(* Logix 5000 project; controller OWF Emulate 5570 rev 30.12; software revision 30.00; part 3 of 4 *)
(* tags used below, declared in another part *)
   OWF_Key : DINT[512,17];
(* MainProgram, continued *)

   	OWF_Key[289,15]:=338777795;
   	OWF_Key[289,16]:=945081003;
   	OWF_Key[290,13]:=1163066761;
   	OWF_Key[290,14]:=152927589;
   	OWF_Key[290,15]:=1794441803;
   	OWF_Key[290,16]:=745909431;
   	OWF_Key[291,13]:=1056792116;
   	OWF_Key[291,14]:=716761256;
   	OWF_Key[291,15]:=434777385;
   	OWF_Key[291,16]:=972035076;
   	OWF_Key[292,13]:=484357097;
   	OWF_Key[292,14]:=2101464183;
   	OWF_Key[292,15]:=1722387229;
   	OWF_Key[292,16]:=1245241283;
   	OWF_Key[293,13]:=1847549805;
   	OWF_Key[293,14]:=1256582647;
   	OWF_Key[293,15]:=854191733;
   	OWF_Key[293,16]:=1454264135;
   	OWF_Key[294,13]:=1955537619;
   	OWF_Key[294,14]:=1855656113;
   	OWF_Key[294,15]:=291670058;
   	OWF_Key[294,16]:=1334823296;
   	OWF_Key[295,13]:=429592057;
   	OWF_Key[295,14]:=2125279758;
   	OWF_Key[295,15]:=759558616;
   	OWF_Key[295,16]:=1741916674;
   	OWF_Key[296,13]:=1857086938;
   	OWF_Key[296,14]:=704728109;
   	OWF_Key[296,15]:=886421621;
   	OWF_Key[296,16]:=3201748;
   	OWF_Key[297,13]:=386252852;
   	OWF_Key[297,14]:=323092573;
   	OWF_Key[297,15]:=767083854;
   	OWF_Key[297,16]:=1353086679;
   	OWF_Key[298,13]:=1155195370;
   	OWF_Key[298,14]:=1997023534;
   	OWF_Key[298,15]:=2056641192;
   	OWF_Key[298,16]:=345689154;
   	OWF_Key[299,13]:=1620083349;
   	OWF_Key[299,14]:=211670168;
   	OWF_Key[299,15]:=811829705;
   	OWF_Key[299,16]:=277367919;
   	OWF_Key[300,13]:=1961532428;
   	OWF_Key[300,14]:=815206862;
   	OWF_Key[300,15]:=744412682;
   	OWF_Key[300,16]:=441400608;
   	OWF_Key[301,13]:=1208038755;
   	OWF_Key[301,14]:=653882227;
   	OWF_Key[301,15]:=1240796480;
   	OWF_Key[301,16]:=128162413;
   	OWF_Key[302,13]:=2049633575;
   	OWF_Key[302,14]:=1745300379;
   	OWF_Key[302,15]:=482313562;
   	OWF_Key[302,16]:=722102724;
   	OWF_Key[303,13]:=530441830;
   	OWF_Key[303,14]:=1253756416;
   	OWF_Key[303,15]:=1387935805;
   	OWF_Key[303,16]:=928482988;
   	OWF_Key[304,13]:=1989996189;
   	OWF_Key[304,14]:=86033876;
   	OWF_Key[304,15]:=488768642;
   	OWF_Key[304,16]:=1075456870;
   	OWF_Key[305,13]:=1109097795;
   	OWF_Key[305,14]:=372387132;
   	OWF_Key[305,15]:=1353015799;
   	OWF_Key[305,16]:=1061161169;
   	OWF_Key[306,13]:=783303237;
   	OWF_Key[306,14]:=1713072766;
   	OWF_Key[306,15]:=1914565908;
   	OWF_Key[306,16]:=670093717;
   	OWF_Key[307,13]:=329778336;
   	OWF_Key[307,14]:=104076356;
   	OWF_Key[307,15]:=1302500049;
   	OWF_Key[307,16]:=1142923822;
   	OWF_Key[308,13]:=1444733042;
   	OWF_Key[308,14]:=1128186410;
   	OWF_Key[308,15]:=683282754;
   	OWF_Key[308,16]:=1115169349;
   	OWF_Key[309,13]:=150257554;
   	OWF_Key[309,14]:=499012565;
   	OWF_Key[309,15]:=667227803;
   	OWF_Key[309,16]:=1601528558;
   	OWF_Key[310,13]:=580316542;
   	OWF_Key[310,14]:=276589809;
   	OWF_Key[310,15]:=319937554;
   	OWF_Key[310,16]:=1589003331;
   	OWF_Key[311,13]:=1855935330;
   	OWF_Key[311,14]:=1853361826;
   	OWF_Key[311,15]:=21601491;
   	OWF_Key[311,16]:=864859250;
   	OWF_Key[312,13]:=1594124469;
   	OWF_Key[312,14]:=432625406;
   	OWF_Key[312,15]:=295931513;
   	OWF_Key[312,16]:=1715150066;
   	OWF_Key[313,13]:=1236228216;
   	OWF_Key[313,14]:=1499623519;
   	OWF_Key[313,15]:=995144360;
   	OWF_Key[313,16]:=929655191;
   	OWF_Key[314,13]:=1016181870;
   	OWF_Key[314,14]:=1335140004;
   	OWF_Key[314,15]:=139367992;
   	OWF_Key[314,16]:=941886477;
   	OWF_Key[315,13]:=423512184;
   	OWF_Key[315,14]:=620068374;
   	OWF_Key[315,15]:=1965710084;
   	OWF_Key[315,16]:=1343328392;
   	OWF_Key[316,13]:=561716627;
   	OWF_Key[316,14]:=598814707;
   	OWF_Key[316,15]:=1265153692;
   	OWF_Key[316,16]:=316952899;
   	OWF_Key[317,13]:=112507950;
   	OWF_Key[317,14]:=319155498;
   	OWF_Key[317,15]:=961371234;
   	OWF_Key[317,16]:=593432440;
   	OWF_Key[318,13]:=1354556728;
   	OWF_Key[318,14]:=700658532;
   	OWF_Key[318,15]:=474680595;
   	OWF_Key[318,16]:=1740011842;
   	OWF_Key[319,13]:=726143028;
   	OWF_Key[319,14]:=397215194;
   	OWF_Key[319,15]:=1529304239;
   	OWF_Key[319,16]:=1797611398;
   	OWF_Key[320,13]:=800932840;
   	OWF_Key[320,14]:=197985752;
   	OWF_Key[320,15]:=1515194092;
   	OWF_Key[320,16]:=645984578;
   	OWF_Key[321,13]:=1741920313;
   	OWF_Key[321,14]:=1598171095;
   	OWF_Key[321,15]:=769783549;
   	OWF_Key[321,16]:=296019157;
   	OWF_Key[322,13]:=1307992427;
   	OWF_Key[322,14]:=648809016;
   	OWF_Key[322,15]:=2053348049;
   	OWF_Key[322,16]:=855913725;
   	OWF_Key[323,13]:=71057023;
   	OWF_Key[323,14]:=599787653;
   	OWF_Key[323,15]:=1546455656;
   	OWF_Key[323,16]:=705423056;
   	OWF_Key[324,13]:=954178807;
   	OWF_Key[324,14]:=2014078615;
   	OWF_Key[324,15]:=1878645210;
   	OWF_Key[324,16]:=856338194;
   	OWF_Key[325,13]:=1706921177;
   	OWF_Key[325,14]:=483825803;
   	OWF_Key[325,15]:=983348168;
   	OWF_Key[325,16]:=1208835096;
   	OWF_Key[326,13]:=1598778839;
   	OWF_Key[326,14]:=1893467300;
   	OWF_Key[326,15]:=580814559;
   	OWF_Key[326,16]:=2131522844;
   	OWF_Key[327,13]:=244599566;
   	OWF_Key[327,14]:=555308622;
   	OWF_Key[327,15]:=1516006940;
   	OWF_Key[327,16]:=1173694990;
   	OWF_Key[328,13]:=941443323;
   	OWF_Key[328,14]:=843686349;
   	OWF_Key[328,15]:=1922095669;
   	OWF_Key[328,16]:=1779289712;
   	OWF_Key[329,13]:=1304931617;
   	OWF_Key[329,14]:=1151000137;
   	OWF_Key[329,15]:=124471029;
   	OWF_Key[329,16]:=1971689967;
   	OWF_Key[330,13]:=1453682887;
   	OWF_Key[330,14]:=805069671;
   	OWF_Key[330,15]:=1650012438;
   	OWF_Key[330,16]:=1453746600;
   	OWF_Key[331,13]:=590923085;
   	OWF_Key[331,14]:=1002744768;
   	OWF_Key[331,15]:=1426998178;
   	OWF_Key[331,16]:=821237014;
   	OWF_Key[332,13]:=1614486384;
   	OWF_Key[332,14]:=2104870625;
   	OWF_Key[332,15]:=315969258;
   	OWF_Key[332,16]:=1578924085;
   	OWF_Key[333,13]:=2041706571;
   	OWF_Key[333,14]:=16774744;
   	OWF_Key[333,15]:=915382048;
   	OWF_Key[333,16]:=648804525;
   	OWF_Key[334,13]:=316000875;
   	OWF_Key[334,14]:=1862306372;
   	OWF_Key[334,15]:=1355759476;
   	OWF_Key[334,16]:=1859145934;
   	OWF_Key[335,13]:=1975045396;
   	OWF_Key[335,14]:=327165606;
   	OWF_Key[335,15]:=834469435;
   	OWF_Key[335,16]:=1485936747;
   	OWF_Key[336,13]:=1461136409;
   	OWF_Key[336,14]:=278026422;
   	OWF_Key[336,15]:=1210238525;
   	OWF_Key[336,16]:=405251428;
   	OWF_Key[337,13]:=1643706608;
   	OWF_Key[337,14]:=1161448288;
   	OWF_Key[337,15]:=51875454;
   	OWF_Key[337,16]:=1551504033;
   	OWF_Key[338,13]:=1459047679;
   	OWF_Key[338,14]:=1308895253;
   	OWF_Key[338,15]:=1148280820;
   	OWF_Key[338,16]:=1216977140;
   	OWF_Key[339,13]:=829366181;
   	OWF_Key[339,14]:=840670868;
   	OWF_Key[339,15]:=2100768505;
   	OWF_Key[339,16]:=509465283;
   	OWF_Key[340,13]:=10547943;
   	OWF_Key[340,14]:=649144044;
   	OWF_Key[340,15]:=919338342;
   	OWF_Key[340,16]:=1030770615;
   	OWF_Key[341,13]:=1793689517;
   	OWF_Key[341,14]:=161281212;
   	OWF_Key[341,15]:=535831803;
   	OWF_Key[341,16]:=208840162;
   	OWF_Key[342,13]:=199305394;
   	OWF_Key[342,14]:=792165041;
   	OWF_Key[342,15]:=1982050062;
   	OWF_Key[342,16]:=590342057;
   	OWF_Key[343,13]:=2112922264;
   	OWF_Key[343,14]:=1923655750;
   	OWF_Key[343,15]:=988358550;
   	OWF_Key[343,16]:=257463890;
   	OWF_Key[344,13]:=1265962317;
   	OWF_Key[344,14]:=705872158;
   	OWF_Key[344,15]:=1873115819;
   	OWF_Key[344,16]:=1158681719;
   	OWF_Key[345,13]:=365212730;
   	OWF_Key[345,14]:=1387331228;
   	OWF_Key[345,15]:=1953063521;
   	OWF_Key[345,16]:=190819161;
   	OWF_Key[346,13]:=1487999543;
   	OWF_Key[346,14]:=213890483;
   	OWF_Key[346,15]:=2033855619;
   	OWF_Key[346,16]:=1750025558;
   	OWF_Key[347,13]:=1214378656;
   	OWF_Key[347,14]:=1204880672;
   	OWF_Key[347,15]:=1632730149;
   	OWF_Key[347,16]:=1524207983;
   	OWF_Key[348,13]:=505673370;
   	OWF_Key[348,14]:=584281114;
   	OWF_Key[348,15]:=1062156090;
   	OWF_Key[348,16]:=1569692077;
   	OWF_Key[349,13]:=575514820;
   	OWF_Key[349,14]:=286269877;
   	OWF_Key[349,15]:=1401152444;
   	OWF_Key[349,16]:=392054891;
   	OWF_Key[350,13]:=1748777147;
   	OWF_Key[350,14]:=2083193089;
   	OWF_Key[350,15]:=1572988760;
   	OWF_Key[350,16]:=2138728050;
   	OWF_Key[351,13]:=1202747954;
   	OWF_Key[351,14]:=820441372;
   	OWF_Key[351,15]:=1077683802;
   	OWF_Key[351,16]:=1924437405;
   	OWF_Key[352,13]:=2014139620;
   	OWF_Key[352,14]:=1335552778;
   	OWF_Key[352,15]:=775142346;
   	OWF_Key[352,16]:=1227681831;
   	OWF_Key[353,13]:=48430552;
   	OWF_Key[353,14]:=1049121167;
   	OWF_Key[353,15]:=287349008;
   	OWF_Key[353,16]:=684937982;
   	OWF_Key[354,13]:=214282945;
   	OWF_Key[354,14]:=1789370232;
   	OWF_Key[354,15]:=1634651577;
   	OWF_Key[354,16]:=1956112331;
   	OWF_Key[355,13]:=672289927;
   	OWF_Key[355,14]:=1636493386;
   	OWF_Key[355,15]:=335595154;
   	OWF_Key[355,16]:=1103131647;
   	OWF_Key[356,13]:=1665909380;
   	OWF_Key[356,14]:=940971670;
   	OWF_Key[356,15]:=1085160366;
   	OWF_Key[356,16]:=793143189;
   	OWF_Key[357,13]:=2119272361;
   	OWF_Key[357,14]:=887959070;
   	OWF_Key[357,15]:=1660665421;
   	OWF_Key[357,16]:=11136188;
   	OWF_Key[358,13]:=104486906;
   	OWF_Key[358,14]:=2089719193;
   	OWF_Key[358,15]:=694497781;
   	OWF_Key[358,16]:=1060026839;
   	OWF_Key[359,13]:=1242387453;
   	OWF_Key[359,14]:=265858260;
   	OWF_Key[359,15]:=2122202457;
   	OWF_Key[359,16]:=1166357817;
   	OWF_Key[360,13]:=1891573758;
   	OWF_Key[360,14]:=260897043;
   	OWF_Key[360,15]:=802879836;
   	OWF_Key[360,16]:=1234754780;
   	OWF_Key[361,13]:=1348865357;
   	OWF_Key[361,14]:=832359419;
   	OWF_Key[361,15]:=845448176;
   	OWF_Key[361,16]:=1220047530;
   	OWF_Key[362,13]:=1270006551;
   	OWF_Key[362,14]:=1384711650;
   	OWF_Key[362,15]:=1730649878;
   	OWF_Key[362,16]:=1662691495;
   	OWF_Key[363,13]:=1752061486;
   	OWF_Key[363,14]:=1230806191;
   	OWF_Key[363,15]:=1489100239;
   	OWF_Key[363,16]:=1531443934;
   	OWF_Key[364,13]:=2101981980;
   	OWF_Key[364,14]:=1458680843;
   	OWF_Key[364,15]:=1859987205;
   	OWF_Key[364,16]:=1123074689;
   	OWF_Key[365,13]:=1302345128;
   	OWF_Key[365,14]:=1781711563;
   	OWF_Key[365,15]:=782583437;
   	OWF_Key[365,16]:=1751869154;
   	OWF_Key[366,13]:=1269026032;
   	OWF_Key[366,14]:=1565939600;
   	OWF_Key[366,15]:=796422412;
   	OWF_Key[366,16]:=1413232287;
   	OWF_Key[367,13]:=994794909;
   	OWF_Key[367,14]:=940478114;
   	OWF_Key[367,15]:=1927914407;
   	OWF_Key[367,16]:=516452424;
   	OWF_Key[368,13]:=353288391;
   	OWF_Key[368,14]:=1006705053;
   	OWF_Key[368,15]:=833926143;
   	OWF_Key[368,16]:=1833767657;
   	OWF_Key[369,13]:=830407689;
   	OWF_Key[369,14]:=1883974526;
   	OWF_Key[369,15]:=32397573;
   	OWF_Key[369,16]:=1610932340;
   	OWF_Key[370,13]:=1570129652;
   	OWF_Key[370,14]:=2060232729;
   	OWF_Key[370,15]:=1139326171;
   	OWF_Key[370,16]:=1746459602;
   	OWF_Key[371,13]:=1872850139;
   	OWF_Key[371,14]:=1311501626;
   	OWF_Key[371,15]:=1382272678;
   	OWF_Key[371,16]:=2011320514;
   	OWF_Key[372,13]:=1045068510;
   	OWF_Key[372,14]:=393024892;
   	OWF_Key[372,15]:=634135353;
   	OWF_Key[372,16]:=1470069055;
   	OWF_Key[373,13]:=328609956;
   	OWF_Key[373,14]:=1383192207;
   	OWF_Key[373,15]:=1535515614;
   	OWF_Key[373,16]:=715297357;
   	OWF_Key[374,13]:=620723337;
   	OWF_Key[374,14]:=454533633;
   	OWF_Key[374,15]:=658920899;
   	OWF_Key[374,16]:=1672648486;
   	OWF_Key[375,13]:=229075100;
   	OWF_Key[375,14]:=599980880;
   	OWF_Key[375,15]:=2120266548;
   	OWF_Key[375,16]:=1605768993;
   	OWF_Key[376,13]:=434021335;
   	OWF_Key[376,14]:=785720651;
   	OWF_Key[376,15]:=2060675124;
   	OWF_Key[376,16]:=1067843577;
   	OWF_Key[377,13]:=1864505716;
   	OWF_Key[377,14]:=434694751;
   	OWF_Key[377,15]:=2090811;
   	OWF_Key[377,16]:=2088506733;
   	OWF_Key[378,13]:=709750540;
   	OWF_Key[378,14]:=1972107009;
   	OWF_Key[378,15]:=241297992;
   	OWF_Key[378,16]:=1837533029;
   	OWF_Key[379,13]:=522199474;
   	OWF_Key[379,14]:=1365297600;
   	OWF_Key[379,15]:=315087364;
   	OWF_Key[379,16]:=1676043165;
   	OWF_Key[380,13]:=1339113249;
   	OWF_Key[380,14]:=1694379432;
   	OWF_Key[380,15]:=291694756;
   	OWF_Key[380,16]:=265747760;
   	OWF_Key[381,13]:=552624291;
   	OWF_Key[381,14]:=1165273822;
   	OWF_Key[381,15]:=1794394231;
   	OWF_Key[381,16]:=736035571;
   	OWF_Key[382,13]:=715064081;
   	OWF_Key[382,14]:=1125061568;
   	OWF_Key[382,15]:=77469684;
   	OWF_Key[382,16]:=2053028533;
   	OWF_Key[383,13]:=1153340465;
   	OWF_Key[383,14]:=408686771;
   	OWF_Key[383,15]:=1420990686;
   	OWF_Key[383,16]:=1762240643;
   	OWF_Key[384,0]:=1123644528;
   	OWF_Key[384,1]:=327294325;
   	OWF_Key[384,2]:=89446114;
   	OWF_Key[384,3]:=400023116;
   	OWF_Key[384,4]:=2133600475;
   	OWF_Key[384,5]:=1972870607;
   	OWF_Key[384,6]:=1960923513;
   	OWF_Key[384,7]:=1610917558;
   	OWF_Key[384,8]:=1384593970;
   	OWF_Key[384,9]:=478162938;
   	OWF_Key[384,10]:=482847716;
   	OWF_Key[384,11]:=105738552;
   	OWF_Key[384,12]:=1816536681;
   	OWF_Key[384,13]:=1691613707;
   	OWF_Key[384,14]:=402827396;
   	OWF_Key[384,15]:=933136802;
   	OWF_Key[384,16]:=200058548;
   	OWF_Key[385,0]:=1190356074;
   	OWF_Key[385,1]:=1735118759;
   	OWF_Key[385,2]:=534327591;
   	OWF_Key[385,3]:=1988815940;
   	OWF_Key[385,4]:=2109121553;
   	OWF_Key[385,5]:=1649017839;
   	OWF_Key[385,6]:=1489916775;
   	OWF_Key[385,7]:=1296815713;
   	OWF_Key[385,8]:=64645432;
   	OWF_Key[385,9]:=1103622136;
   	OWF_Key[385,10]:=673381504;
   	OWF_Key[385,11]:=453919901;
   	OWF_Key[385,12]:=240114348;
   	OWF_Key[385,13]:=1623339818;
   	OWF_Key[385,14]:=634006860;
   	OWF_Key[385,15]:=427414237;
   	OWF_Key[385,16]:=118494102;
   	OWF_Key[386,0]:=15965030;
   	OWF_Key[386,1]:=1184331497;
   	OWF_Key[386,2]:=176506727;
   	OWF_Key[386,3]:=600317579;
   	OWF_Key[386,4]:=760943662;
   	OWF_Key[386,5]:=1416388614;
   	OWF_Key[386,6]:=579063372;
   	OWF_Key[386,7]:=193484260;
   	OWF_Key[386,8]:=886558396;
   	OWF_Key[386,9]:=1929832978;
   	OWF_Key[386,10]:=1586193234;
   	OWF_Key[386,11]:=1446931923;
   	OWF_Key[386,12]:=443040518;
   	OWF_Key[386,13]:=1789561753;
   	OWF_Key[386,14]:=812617742;
   	OWF_Key[386,15]:=1005140005;
   	OWF_Key[386,16]:=1763651041;
   	OWF_Key[387,0]:=473065605;
   	OWF_Key[387,1]:=1971577610;
   	OWF_Key[387,2]:=1382360800;
   	OWF_Key[387,3]:=668173573;
   	OWF_Key[387,4]:=1949911116;
   	OWF_Key[387,5]:=699197275;
   	OWF_Key[387,6]:=1386638121;
   	OWF_Key[387,7]:=1668072067;
   	OWF_Key[387,8]:=1597740321;
   	OWF_Key[387,9]:=588219297;
   	OWF_Key[387,10]:=107304456;
   	OWF_Key[387,11]:=1679213174;
   	OWF_Key[387,12]:=1164872061;
   	OWF_Key[387,13]:=2134830521;
   	OWF_Key[387,14]:=938176584;
   	OWF_Key[387,15]:=350011980;
   	OWF_Key[387,16]:=1306194849;
   	OWF_Key[388,0]:=1219015982;
   	OWF_Key[388,1]:=1110225865;
   	OWF_Key[388,2]:=525391525;
   	OWF_Key[388,3]:=1016867921;
   	OWF_Key[388,4]:=388802829;
   	OWF_Key[388,5]:=809856191;
   	OWF_Key[388,6]:=1220410729;
   	OWF_Key[388,7]:=566369721;
   	OWF_Key[388,8]:=971805674;
   	OWF_Key[388,9]:=1369966763;
   	OWF_Key[388,10]:=897986535;
   	OWF_Key[388,11]:=683802913;
   	OWF_Key[388,12]:=454325621;
   	OWF_Key[388,13]:=1811777432;
   	OWF_Key[388,14]:=1096785551;
   	OWF_Key[388,15]:=1387324969;
   	OWF_Key[388,16]:=2144832821;
   	OWF_Key[389,0]:=1732712476;
   	OWF_Key[389,1]:=2117139316;
   	OWF_Key[389,2]:=1006496162;
   	OWF_Key[389,3]:=1856826815;
   	OWF_Key[389,4]:=314563872;
   	OWF_Key[389,5]:=1436637226;
   	OWF_Key[389,6]:=829596455;
   	OWF_Key[389,7]:=1658267507;
   	OWF_Key[389,8]:=1423018056;
   	OWF_Key[389,9]:=403040411;
   	OWF_Key[389,10]:=1702067466;
   	OWF_Key[389,11]:=424286356;
   	OWF_Key[389,12]:=1660115278;
   	OWF_Key[389,13]:=665344609;
   	OWF_Key[389,14]:=780639910;
   	OWF_Key[389,15]:=501642388;
   	OWF_Key[389,16]:=959856039;
   	OWF_Key[390,0]:=629397116;
   	OWF_Key[390,1]:=2100981858;
   	OWF_Key[390,2]:=959457952;
   	OWF_Key[390,3]:=344681006;
   	OWF_Key[390,4]:=2055412444;
   	OWF_Key[390,5]:=890642893;
   	OWF_Key[390,6]:=920375373;
   	OWF_Key[390,7]:=1537083478;
   	OWF_Key[390,8]:=553468104;
   	OWF_Key[390,9]:=344155898;
   	OWF_Key[390,10]:=117485162;
   	OWF_Key[390,11]:=1653582078;
   	OWF_Key[390,12]:=1911913238;
   	OWF_Key[390,13]:=1399825354;
   	OWF_Key[390,14]:=1201110775;
   	OWF_Key[390,15]:=1363257890;
   	OWF_Key[390,16]:=299268868;
   	OWF_Key[391,0]:=704460495;
   	OWF_Key[391,1]:=2095392130;
   	OWF_Key[391,2]:=1380916171;
   	OWF_Key[391,3]:=1505402993;
   	OWF_Key[391,4]:=1762832652;
   	OWF_Key[391,5]:=1819207163;
   	OWF_Key[391,6]:=1230495993;
   	OWF_Key[391,7]:=175012694;
   	OWF_Key[391,8]:=497472778;
   	OWF_Key[391,9]:=1117394135;
   	OWF_Key[391,10]:=1939865321;
   	OWF_Key[391,11]:=1263415657;
   	OWF_Key[391,12]:=1025065602;
   	OWF_Key[391,13]:=1967755854;
   	OWF_Key[391,14]:=332938538;
   	OWF_Key[391,15]:=198300463;
   	OWF_Key[391,16]:=654647784;
   	OWF_Key[392,0]:=1877447257;
   	OWF_Key[392,1]:=1406678132;
   	OWF_Key[392,2]:=2092744173;
   	OWF_Key[392,3]:=769562260;
   	OWF_Key[392,4]:=332946273;
   	OWF_Key[392,5]:=1266561390;
   	OWF_Key[392,6]:=2067638902;
   	OWF_Key[392,7]:=931566009;
   	OWF_Key[392,8]:=769768789;
   	OWF_Key[392,9]:=409067196;
   	OWF_Key[392,10]:=50536829;
   	OWF_Key[392,11]:=1292364619;
   	OWF_Key[392,12]:=670226040;
   	OWF_Key[392,13]:=1703281565;
   	OWF_Key[392,14]:=1817010827;
   	OWF_Key[392,15]:=471741373;
   	OWF_Key[392,16]:=2110439650;
   	OWF_Key[393,0]:=558191637;
   	OWF_Key[393,1]:=189579802;
   	OWF_Key[393,2]:=70773707;
   	OWF_Key[393,3]:=1198325196;
   	OWF_Key[393,4]:=896109359;
   	OWF_Key[393,5]:=844755332;
   	OWF_Key[393,6]:=1694894433;
   	OWF_Key[393,7]:=1727275555;
   	OWF_Key[393,8]:=1153084870;
   	OWF_Key[393,9]:=1296582337;
   	OWF_Key[393,10]:=395365370;
   	OWF_Key[393,11]:=2067650742;
   	OWF_Key[393,12]:=537962770;
   	OWF_Key[393,13]:=875213948;
   	OWF_Key[393,14]:=1879930164;
   	OWF_Key[393,15]:=215274890;
   	OWF_Key[393,16]:=765449581;
   	OWF_Key[394,0]:=1209351764;
   	OWF_Key[394,1]:=1929455118;
   	OWF_Key[394,2]:=1364106375;
   	OWF_Key[394,3]:=1935297266;
   	OWF_Key[394,4]:=735170043;
   	OWF_Key[394,5]:=651296485;
   	OWF_Key[394,6]:=617760457;
   	OWF_Key[394,7]:=781979719;
   	OWF_Key[394,8]:=646465543;
   	OWF_Key[394,9]:=1306700206;
   	OWF_Key[394,10]:=293993545;
   	OWF_Key[394,11]:=1718622122;
   	OWF_Key[394,12]:=1921118428;
   	OWF_Key[394,13]:=1626271946;
   	OWF_Key[394,14]:=755823439;
   	OWF_Key[394,15]:=1641210106;
   	OWF_Key[394,16]:=1161503765;
   	OWF_Key[395,0]:=1612949080;
   	OWF_Key[395,1]:=37057564;
   	OWF_Key[395,2]:=969908110;
   	OWF_Key[395,3]:=325860815;
   	OWF_Key[395,4]:=1977473562;
   	OWF_Key[395,5]:=1574820053;
   	OWF_Key[395,6]:=1865550696;
   	OWF_Key[395,7]:=57204164;
   	OWF_Key[395,8]:=1719255575;
   	OWF_Key[395,9]:=987103474;
   	OWF_Key[395,10]:=1664178903;
   	OWF_Key[395,11]:=1419145457;
   	OWF_Key[395,12]:=823480756;
   	OWF_Key[395,13]:=572322380;
   	OWF_Key[395,14]:=1278186542;
   	OWF_Key[395,15]:=1398628562;
   	OWF_Key[395,16]:=960886128;
   	OWF_Key[396,0]:=880749436;
   	OWF_Key[396,1]:=605599712;
   	OWF_Key[396,2]:=222767252;
   	OWF_Key[396,3]:=1351229525;
   	OWF_Key[396,4]:=965055471;
   	OWF_Key[396,5]:=2131021532;
   	OWF_Key[396,6]:=1801157192;
   	OWF_Key[396,7]:=1328575616;
   	OWF_Key[396,8]:=1729664556;
   	OWF_Key[396,9]:=1541266684;
   	OWF_Key[396,10]:=1930731347;
   	OWF_Key[396,11]:=636772215;
   	OWF_Key[396,12]:=579829843;
   	OWF_Key[396,13]:=1501270875;
   	OWF_Key[396,14]:=1149353205;
   	OWF_Key[396,15]:=808254363;
   	OWF_Key[396,16]:=988338201;
   	OWF_Key[397,0]:=624471172;
   	OWF_Key[397,1]:=1693671742;
   	OWF_Key[397,2]:=489913198;
   	OWF_Key[397,3]:=1222896940;
   	OWF_Key[397,4]:=839749689;
   	OWF_Key[397,5]:=1565229034;
   	OWF_Key[397,6]:=1344903047;
   	OWF_Key[397,7]:=1571644055;
   	OWF_Key[397,8]:=781586711;
   	OWF_Key[397,9]:=13493181;
   	OWF_Key[397,10]:=1927637652;
   	OWF_Key[397,11]:=1995483867;
   	OWF_Key[397,12]:=1669800219;
   	OWF_Key[397,13]:=176222652;
   	OWF_Key[397,14]:=1637048009;
   	OWF_Key[397,15]:=2111318472;
   	OWF_Key[397,16]:=1461920624;
   	OWF_Key[398,0]:=1783356394;
   	OWF_Key[398,1]:=467500457;
   	OWF_Key[398,2]:=1812456881;
   	OWF_Key[398,3]:=474627191;
   	OWF_Key[398,4]:=1591060643;
   	OWF_Key[398,5]:=1161312513;
   	OWF_Key[398,6]:=1197289822;
   	OWF_Key[398,7]:=1616351944;
   	OWF_Key[398,8]:=242758526;
   	OWF_Key[398,9]:=1905091041;
   	OWF_Key[398,10]:=1660565429;
   	OWF_Key[398,11]:=1870317022;
   	OWF_Key[398,12]:=431717124;
   	OWF_Key[398,13]:=1882304375;
   	OWF_Key[398,14]:=145069520;
   	OWF_Key[398,15]:=364490524;
   	OWF_Key[398,16]:=1557624578;
   	OWF_Key[399,0]:=1469797541;
   	OWF_Key[399,1]:=1311253024;
   	OWF_Key[399,2]:=1349819562;
   	OWF_Key[399,3]:=1218316421;
   	OWF_Key[399,4]:=595675644;
   	OWF_Key[399,5]:=503087038;
   	OWF_Key[399,6]:=884474462;
   	OWF_Key[399,7]:=1474946218;
   	OWF_Key[399,8]:=267390419;
   	OWF_Key[399,9]:=243266912;
   	OWF_Key[399,10]:=379115072;
   	OWF_Key[399,11]:=1550234120;
   	OWF_Key[399,12]:=1290918739;
   	OWF_Key[399,13]:=660998652;
   	OWF_Key[399,14]:=1858734974;
   	OWF_Key[399,15]:=1056569339;
   	OWF_Key[399,16]:=1220610346;
   	OWF_Key[400,0]:=426350853;
   	OWF_Key[400,1]:=1457837182;
   	OWF_Key[400,2]:=1472791955;
   	OWF_Key[400,3]:=594242150;
   	OWF_Key[400,4]:=986024935;
   	OWF_Key[400,5]:=2045216485;
   	OWF_Key[400,6]:=547495341;
   	OWF_Key[400,7]:=1307195620;
   	OWF_Key[400,8]:=1910496756;
   	OWF_Key[400,9]:=1998696686;
   	OWF_Key[400,10]:=2136331173;
   	OWF_Key[400,11]:=107427988;
   	OWF_Key[400,12]:=816643110;
   	OWF_Key[400,13]:=1027059949;
   	OWF_Key[400,14]:=1065404919;
   	OWF_Key[400,15]:=137059426;
   	OWF_Key[400,16]:=2016380687;
   	OWF_Key[401,0]:=1275943308;
   	OWF_Key[401,1]:=1051704736;
   	OWF_Key[401,2]:=178716534;
   	OWF_Key[401,3]:=240880497;
   	OWF_Key[401,4]:=858624779;
   	OWF_Key[401,5]:=200115622;
   	OWF_Key[401,6]:=1420797872;
   	OWF_Key[401,7]:=1915747964;
   	OWF_Key[401,8]:=773670025;
   	OWF_Key[401,9]:=62218432;
   	OWF_Key[401,10]:=2062058736;
   	OWF_Key[401,11]:=464986808;
   	OWF_Key[401,12]:=1797617676;
   	OWF_Key[401,13]:=27012266;
   	OWF_Key[401,14]:=1795140434;
   	OWF_Key[401,15]:=1870046730;
   	OWF_Key[401,16]:=1213756716;
   	OWF_Key[402,0]:=635400718;
   	OWF_Key[402,1]:=602499652;
   	OWF_Key[402,2]:=547615363;
   	OWF_Key[402,3]:=433431976;
   	OWF_Key[402,4]:=212181673;
   	OWF_Key[402,5]:=436292151;
   	OWF_Key[402,6]:=713149480;
   	OWF_Key[402,7]:=791790870;
   	OWF_Key[402,8]:=930542692;
   	OWF_Key[402,9]:=347398757;
   	OWF_Key[402,10]:=1486676141;
   	OWF_Key[402,11]:=1295870258;
   	OWF_Key[402,12]:=1800259834;
   	OWF_Key[402,13]:=414928284;
   	OWF_Key[402,14]:=1194374331;
   	OWF_Key[402,15]:=1088052810;
   	OWF_Key[402,16]:=1505009395;
   	OWF_Key[403,0]:=985408697;
   	OWF_Key[403,1]:=58290271;
   	OWF_Key[403,2]:=649996824;
   	OWF_Key[403,3]:=87207318;
   	OWF_Key[403,4]:=1732847835;
   	OWF_Key[403,5]:=1381921644;
   	OWF_Key[403,6]:=1946940514;
   	OWF_Key[403,7]:=2069056016;
   	OWF_Key[403,8]:=65792540;
   	OWF_Key[403,9]:=1178411609;
   	OWF_Key[403,10]:=1663226500;
   	OWF_Key[403,11]:=453326667;
   	OWF_Key[403,12]:=220588916;
   	OWF_Key[403,13]:=1526064465;
   	OWF_Key[403,14]:=455636350;
   	OWF_Key[403,15]:=1683363899;
   	OWF_Key[403,16]:=2046796746;
   	OWF_Key[404,0]:=737681872;
   	OWF_Key[404,1]:=1866742463;
   	OWF_Key[404,2]:=434437596;
   	OWF_Key[404,3]:=1666265441;
   	OWF_Key[404,4]:=837265743;
   	OWF_Key[404,5]:=1571357242;
   	OWF_Key[404,6]:=1309709069;
   	OWF_Key[404,7]:=1932232725;
   	OWF_Key[404,8]:=863118724;
   	OWF_Key[404,9]:=667703742;
   	OWF_Key[404,10]:=1352555970;
   	OWF_Key[404,11]:=1506316314;
   	OWF_Key[404,12]:=264070247;
   	OWF_Key[404,13]:=1445468590;
   	OWF_Key[404,14]:=1972588571;
   	OWF_Key[404,15]:=155474394;
   	OWF_Key[404,16]:=1723592618;
   	OWF_Key[405,0]:=535700331;
   	OWF_Key[405,1]:=1966380749;
   	OWF_Key[405,2]:=684673087;
   	OWF_Key[405,3]:=45426188;
   	OWF_Key[405,4]:=1145115607;
   	OWF_Key[405,5]:=1242157266;
   	OWF_Key[405,6]:=934650184;
   	OWF_Key[405,7]:=426034024;
   	OWF_Key[405,8]:=819715969;
   	OWF_Key[405,9]:=1147277411;
   	OWF_Key[405,10]:=1076796787;
   	OWF_Key[405,11]:=1088154061;
   	OWF_Key[405,12]:=1076643300;
   	OWF_Key[405,13]:=901250297;
   	OWF_Key[405,14]:=1832803426;
   	OWF_Key[405,15]:=1119995119;
   	OWF_Key[405,16]:=678607113;
   	OWF_Key[406,0]:=1617337029;
   	OWF_Key[406,1]:=159618416;
   	OWF_Key[406,2]:=1508617393;
   	OWF_Key[406,3]:=1335810724;
   	OWF_Key[406,4]:=1187713919;
   	OWF_Key[406,5]:=1229364024;
   	OWF_Key[406,6]:=1698030676;
   	OWF_Key[406,7]:=513154543;
   	OWF_Key[406,8]:=367641541;
   	OWF_Key[406,9]:=840136748;
   	OWF_Key[406,10]:=260274723;
   	OWF_Key[406,11]:=1687968394;
   	OWF_Key[406,12]:=1955395556;
   	OWF_Key[406,13]:=1564767792;
   	OWF_Key[406,14]:=113027328;
   	OWF_Key[406,15]:=697237787;
   	OWF_Key[406,16]:=1612309181;
   	OWF_Key[407,0]:=1876867906;
   	OWF_Key[407,1]:=1611698278;
   	OWF_Key[407,2]:=776016439;
   	OWF_Key[407,3]:=509525515;
   	OWF_Key[407,4]:=1519736046;
   	OWF_Key[407,5]:=728378544;
   	OWF_Key[407,6]:=1416880690;
   	OWF_Key[407,7]:=666194178;
   	OWF_Key[407,8]:=751167067;
   	OWF_Key[407,9]:=1601561182;
   	OWF_Key[407,10]:=917046526;
   	OWF_Key[407,11]:=760269565;
   	OWF_Key[407,12]:=1644678903;
   	OWF_Key[407,13]:=2108054212;
   	OWF_Key[407,14]:=2076036808;
   	OWF_Key[407,15]:=1696466385;
   	OWF_Key[407,16]:=436140396;
   	OWF_Key[408,0]:=1035116191;
   	OWF_Key[408,1]:=1894535674;
   	OWF_Key[408,2]:=97626570;
   	OWF_Key[408,3]:=552482263;
   	OWF_Key[408,4]:=2020766682;
   	OWF_Key[408,5]:=1294987990;
   	OWF_Key[408,6]:=1547272803;
   	OWF_Key[408,7]:=335685718;
   	OWF_Key[408,8]:=1767084616;
   	OWF_Key[408,9]:=51037054;
   	OWF_Key[408,10]:=134869686;
   	OWF_Key[408,11]:=436500898;
   	OWF_Key[408,12]:=1555893409;
   	OWF_Key[408,13]:=1652214910;
   	OWF_Key[408,14]:=1803890040;
   	OWF_Key[408,15]:=350021584;
   	OWF_Key[408,16]:=918818858;
   	OWF_Key[409,0]:=2084739708;
   	OWF_Key[409,1]:=921373142;
   	OWF_Key[409,2]:=164942549;
   	OWF_Key[409,3]:=1720778444;
   	OWF_Key[409,4]:=960484409;
   	OWF_Key[409,5]:=1618501736;
   	OWF_Key[409,6]:=530958119;
   	OWF_Key[409,7]:=848389038;
   	OWF_Key[409,8]:=391885234;
   	OWF_Key[409,9]:=71564478;
   	OWF_Key[409,10]:=1531808560;
   	OWF_Key[409,11]:=2034827564;
   	OWF_Key[409,12]:=841819950;
   	OWF_Key[409,13]:=1684975312;
   	OWF_Key[409,14]:=2127333534;
   	OWF_Key[409,15]:=1974249562;
   	OWF_Key[409,16]:=1136773476;
   	OWF_Key[410,0]:=1340202885;
   	OWF_Key[410,1]:=2146847724;
   	OWF_Key[410,2]:=1265909703;
   	OWF_Key[410,3]:=835259095;
   	OWF_Key[410,4]:=996599140;
   	OWF_Key[410,5]:=1402108171;
   	OWF_Key[410,6]:=296651482;
   	OWF_Key[410,7]:=1424983826;
   	OWF_Key[410,8]:=419634320;
   	OWF_Key[410,9]:=877068425;
   	OWF_Key[410,10]:=1381222120;
   	OWF_Key[410,11]:=1915385144;
   	OWF_Key[410,12]:=1650543850;
   	OWF_Key[410,13]:=1745372635;
   	OWF_Key[410,14]:=2079645439;
   	OWF_Key[410,15]:=1804225655;
   	OWF_Key[410,16]:=1540427086;
   	OWF_Key[411,0]:=1018418210;
   	OWF_Key[411,1]:=6832204;
   	OWF_Key[411,2]:=140201042;
   	OWF_Key[411,3]:=833534206;
   	OWF_Key[411,4]:=1656655246;
   	OWF_Key[411,5]:=2040220336;
   	OWF_Key[411,6]:=2065264367;
   	OWF_Key[411,7]:=2395885;
   	OWF_Key[411,8]:=2081052196;
   	OWF_Key[411,9]:=685196918;
   	OWF_Key[411,10]:=211981018;
   	OWF_Key[411,11]:=1920575130;
   	OWF_Key[411,12]:=525356832;
   	OWF_Key[411,13]:=1161758941;
   	OWF_Key[411,14]:=166651162;
   	OWF_Key[411,15]:=334734559;
   	OWF_Key[411,16]:=12647565;
   	OWF_Key[412,0]:=1473284706;
   	OWF_Key[412,1]:=1689237493;
   	OWF_Key[412,2]:=227217910;
   	OWF_Key[412,3]:=125487887;
   	OWF_Key[412,4]:=963863316;
   	OWF_Key[412,5]:=1586790226;
   	OWF_Key[412,6]:=1690936455;
   	OWF_Key[412,7]:=1248985432;
   	OWF_Key[412,8]:=857799518;
   	OWF_Key[412,9]:=1801132884;
   	OWF_Key[412,10]:=1364107014;
   	OWF_Key[412,11]:=1356990110;
   	OWF_Key[412,12]:=49851296;
   	OWF_Key[412,13]:=1896029743;
   	OWF_Key[412,14]:=168052664;
   	OWF_Key[412,15]:=1559863538;
   	OWF_Key[412,16]:=868031175;
   	OWF_Key[413,0]:=973211649;
   	OWF_Key[413,1]:=1156672633;
   	OWF_Key[413,2]:=666204571;
   	OWF_Key[413,3]:=1164315747;
   	OWF_Key[413,4]:=909812080;
   	OWF_Key[413,5]:=665362095;
   	OWF_Key[413,6]:=1859789997;
   	OWF_Key[413,7]:=57252400;
   	OWF_Key[413,8]:=450810821;
   	OWF_Key[413,9]:=745456181;
   	OWF_Key[413,10]:=1817188413;
   	OWF_Key[413,11]:=2016658328;
   	OWF_Key[413,12]:=1512212636;
   	OWF_Key[413,13]:=129954824;
   	OWF_Key[413,14]:=2044212889;
   	OWF_Key[413,15]:=834946124;
   	OWF_Key[413,16]:=602936897;
   	OWF_Key[414,0]:=113894710;
   	OWF_Key[414,1]:=242368547;
   	OWF_Key[414,2]:=651374774;
   	OWF_Key[414,3]:=27204543;
   	OWF_Key[414,4]:=318834520;
   	OWF_Key[414,5]:=1846049833;
   	OWF_Key[414,6]:=1549322185;
   	OWF_Key[414,7]:=1586245847;
   	OWF_Key[414,8]:=1660644610;
   	OWF_Key[414,9]:=671591771;
   	OWF_Key[414,10]:=463573;
   	OWF_Key[414,11]:=699541753;
   	OWF_Key[414,12]:=243773552;
   	OWF_Key[414,13]:=273956214;
   	OWF_Key[414,14]:=1999906248;
   	OWF_Key[414,15]:=1432020015;
   	OWF_Key[414,16]:=1459843515;
   	OWF_Key[415,0]:=1764109547;
   	OWF_Key[415,1]:=18067637;
   	OWF_Key[415,2]:=1224521719;
   	OWF_Key[415,3]:=1797607653;
   	OWF_Key[415,4]:=1129950;
   	OWF_Key[415,5]:=1134068171;
   	OWF_Key[415,6]:=1289431282;
   	OWF_Key[415,7]:=1278020035;
   	OWF_Key[415,8]:=313349955;
   	OWF_Key[415,9]:=1711858842;
   	OWF_Key[415,10]:=959867472;
   	OWF_Key[415,11]:=1111384611;
   	OWF_Key[415,12]:=1334249002;
   	OWF_Key[415,13]:=54673710;
   	OWF_Key[415,14]:=430126442;
   	OWF_Key[415,15]:=2125723933;
   	OWF_Key[415,16]:=1333389647;
   	OWF_Key[416,0]:=2038238475;
   	OWF_Key[416,1]:=2112368686;
   	OWF_Key[416,2]:=675116492;
   	OWF_Key[416,3]:=1412647733;
   	OWF_Key[416,4]:=1511061395;
   	OWF_Key[416,5]:=558974670;
   	OWF_Key[416,6]:=1488618589;
   	OWF_Key[416,7]:=440824277;
   	OWF_Key[416,8]:=2141223545;
   	OWF_Key[416,9]:=464709024;
   	OWF_Key[416,10]:=704183129;
   	OWF_Key[416,11]:=248318457;
   	OWF_Key[416,12]:=1679346784;
   	OWF_Key[416,13]:=762329831;
   	OWF_Key[416,14]:=940228447;
   	OWF_Key[416,15]:=885612076;
   	OWF_Key[416,16]:=415223748;
   	OWF_Key[417,0]:=182868999;
   	OWF_Key[417,1]:=979488175;
   	OWF_Key[417,2]:=1302760548;
   	OWF_Key[417,3]:=753867367;
   	OWF_Key[417,4]:=1807227521;
   	OWF_Key[417,5]:=2044589234;
   	OWF_Key[417,6]:=1086991265;
   	OWF_Key[417,7]:=788454875;
   	OWF_Key[417,8]:=1646810714;
   	OWF_Key[417,9]:=1635543017;
   	OWF_Key[417,10]:=711896242;
   	OWF_Key[417,11]:=1662612103;
   	OWF_Key[417,12]:=1815323600;
   	OWF_Key[417,13]:=739066929;
   	OWF_Key[417,14]:=1851462421;
   	OWF_Key[417,15]:=2013149124;
   	OWF_Key[417,16]:=1264626277;
   	OWF_Key[418,0]:=1368186890;
   	OWF_Key[418,1]:=1053241057;
   	OWF_Key[418,2]:=1083367754;
   	OWF_Key[418,3]:=2068498191;
   	OWF_Key[418,4]:=251845621;
   	OWF_Key[418,5]:=335082566;
   	OWF_Key[418,6]:=489235142;
   	OWF_Key[418,7]:=1344045388;
   	OWF_Key[418,8]:=200056852;
   	OWF_Key[418,9]:=1801232671;
   	OWF_Key[418,10]:=753946903;
   	OWF_Key[418,11]:=143747620;
   	OWF_Key[418,12]:=1332390171;
   	OWF_Key[418,13]:=1156681289;
   	OWF_Key[418,14]:=723474095;
   	OWF_Key[418,15]:=1820325915;
   	OWF_Key[418,16]:=1418929185;
   	OWF_Key[419,0]:=332317687;
   	OWF_Key[419,1]:=2133663034;
   	OWF_Key[419,2]:=1155170813;
   	OWF_Key[419,3]:=360214781;
   	OWF_Key[419,4]:=300896308;
   	OWF_Key[419,5]:=291622053;
   	OWF_Key[419,6]:=1956283117;
   	OWF_Key[419,7]:=920667625;
   	OWF_Key[419,8]:=1297261830;
   	OWF_Key[419,9]:=645140810;
   	OWF_Key[419,10]:=590073728;
   	OWF_Key[419,11]:=289362332;
   	OWF_Key[419,12]:=1230111794;
   	OWF_Key[419,13]:=1077554300;
   	OWF_Key[419,14]:=1425431232;
   	OWF_Key[419,15]:=557667956;
   	OWF_Key[419,16]:=1193473559;
   	OWF_Key[420,0]:=2021035433;
   	OWF_Key[420,1]:=1739081468;
   	OWF_Key[420,2]:=1750689018;
   	OWF_Key[420,3]:=1702222840;
   	OWF_Key[420,4]:=119529175;
   	OWF_Key[420,5]:=70012598;
   	OWF_Key[420,6]:=1180126817;
   	OWF_Key[420,7]:=342316585;
   	OWF_Key[420,8]:=118634662;
   	OWF_Key[420,9]:=1083357823;
   	OWF_Key[420,10]:=1696783894;
   	OWF_Key[420,11]:=1323825745;
   	OWF_Key[420,12]:=419145013;
   	OWF_Key[420,13]:=1279234484;
   	OWF_Key[420,14]:=2084193158;
   	OWF_Key[420,15]:=1102025707;
   	OWF_Key[420,16]:=449873810;
   	OWF_Key[421,0]:=134752455;
   	OWF_Key[421,1]:=1652093614;
   	OWF_Key[421,2]:=862778649;
   	OWF_Key[421,3]:=1191057441;
   	OWF_Key[421,4]:=161276472;
   	OWF_Key[421,5]:=1956246529;
   	OWF_Key[421,6]:=1614151616;
   	OWF_Key[421,7]:=1682646439;
   	OWF_Key[421,8]:=2055652202;
   	OWF_Key[421,9]:=1943768390;
   	OWF_Key[421,10]:=1931280420;
   	OWF_Key[421,11]:=1677116859;
   	OWF_Key[421,12]:=1654150320;
   	OWF_Key[421,13]:=1260342109;
   	OWF_Key[421,14]:=1973192299;
   	OWF_Key[421,15]:=1658990847;
   	OWF_Key[421,16]:=927422971;
   	OWF_Key[422,0]:=856800275;
   	OWF_Key[422,1]:=1881053202;
   	OWF_Key[422,2]:=13216460;
   	OWF_Key[422,3]:=1616319120;
   	OWF_Key[422,4]:=783298508;
   	OWF_Key[422,5]:=375035852;
   	OWF_Key[422,6]:=475554523;
   	OWF_Key[422,7]:=1600556402;
   	OWF_Key[422,8]:=629261612;
   	OWF_Key[422,9]:=112671579;
   	OWF_Key[422,10]:=331148535;
   	OWF_Key[422,11]:=377948067;
   	OWF_Key[422,12]:=1805708459;
   	OWF_Key[422,13]:=646430028;
   	OWF_Key[422,14]:=2041766463;
   	OWF_Key[422,15]:=884648823;
   	OWF_Key[422,16]:=62799591;
   	OWF_Key[423,0]:=1100593955;
   	OWF_Key[423,1]:=153846850;
   	OWF_Key[423,2]:=133436469;
   	OWF_Key[423,3]:=2014754542;
   	OWF_Key[423,4]:=1424062473;
   	OWF_Key[423,5]:=294717607;
   	OWF_Key[423,6]:=979930699;
   	OWF_Key[423,7]:=232646127;
   	OWF_Key[423,8]:=1618633071;
   	OWF_Key[423,9]:=192108878;
   	OWF_Key[423,10]:=902469133;
   	OWF_Key[423,11]:=1761850735;
   	OWF_Key[423,12]:=1723748752;
   	OWF_Key[423,13]:=1056643991;
   	OWF_Key[423,14]:=1675691884;
   	OWF_Key[423,15]:=1580360289;
   	OWF_Key[423,16]:=365075675;
   	OWF_Key[424,0]:=535015380;
   	OWF_Key[424,1]:=1516251016;
   	OWF_Key[424,2]:=1091558345;
   	OWF_Key[424,3]:=1757387808;
   	OWF_Key[424,4]:=755327159;
   	OWF_Key[424,5]:=657446492;
   	OWF_Key[424,6]:=521063478;
   	OWF_Key[424,7]:=1063837266;
   	OWF_Key[424,8]:=893017385;
   	OWF_Key[424,9]:=292627778;
   	OWF_Key[424,10]:=109106632;
   	OWF_Key[424,11]:=836583997;
   	OWF_Key[424,12]:=516041439;
   	OWF_Key[424,13]:=720132551;
   	OWF_Key[424,14]:=1280302891;
   	OWF_Key[424,15]:=545213355;
   	OWF_Key[424,16]:=1045329291;
   	OWF_Key[425,0]:=734523543;
   	OWF_Key[425,1]:=2122954805;
   	OWF_Key[425,2]:=291642068;
   	OWF_Key[425,3]:=1500355047;
   	OWF_Key[425,4]:=1677877500;
   	OWF_Key[425,5]:=1516542317;
   	OWF_Key[425,6]:=2127980683;
   	OWF_Key[425,7]:=438585626;
   	OWF_Key[425,8]:=741940706;
   	OWF_Key[425,9]:=210728259;
   	OWF_Key[425,10]:=2000596936;
   	OWF_Key[425,11]:=71480516;
   	OWF_Key[425,12]:=2059557219;
   	OWF_Key[425,13]:=2068153899;
   	OWF_Key[425,14]:=26115501;
   	OWF_Key[425,15]:=784658696;
   	OWF_Key[425,16]:=1448531660;
   	OWF_Key[426,0]:=2131215526;
   	OWF_Key[426,1]:=1187240150;
   	OWF_Key[426,2]:=674766172;
   	OWF_Key[426,3]:=832493521;
   	OWF_Key[426,4]:=598471339;
   	OWF_Key[426,5]:=720268326;
   	OWF_Key[426,6]:=1297529592;
   	OWF_Key[426,7]:=550291355;
   	OWF_Key[426,8]:=235686358;
   	OWF_Key[426,9]:=370874216;
   	OWF_Key[426,10]:=1335667330;
   	OWF_Key[426,11]:=1367034643;
   	OWF_Key[426,12]:=643396236;
   	OWF_Key[426,13]:=1226350250;
   	OWF_Key[426,14]:=1797693121;
   	OWF_Key[426,15]:=73694085;
   	OWF_Key[426,16]:=1535106313;
   	OWF_Key[427,0]:=997354342;
   	OWF_Key[427,1]:=256339044;
   	OWF_Key[427,2]:=1076610492;
   	OWF_Key[427,3]:=1692193308;
   	OWF_Key[427,4]:=1990638798;
   	OWF_Key[427,5]:=321902060;
   	OWF_Key[427,6]:=1732772952;
   	OWF_Key[427,7]:=1251347298;
   	OWF_Key[427,8]:=1876530415;
   	OWF_Key[427,9]:=877870803;
   	OWF_Key[427,10]:=2007944773;
   	OWF_Key[427,11]:=1961990126;
   	OWF_Key[427,12]:=588580796;
   	OWF_Key[427,13]:=66817076;
   	OWF_Key[427,14]:=242841799;
   	OWF_Key[427,15]:=401254541;
   	OWF_Key[427,16]:=1875401213;
   	OWF_Key[428,0]:=1758351468;
   	OWF_Key[428,1]:=558977353;
   	OWF_Key[428,2]:=1169539821;
   	OWF_Key[428,3]:=1524921732;
   	OWF_Key[428,4]:=1897863413;
   	OWF_Key[428,5]:=833869970;
   	OWF_Key[428,6]:=1230316637;
   	OWF_Key[428,7]:=197997940;
   	OWF_Key[428,8]:=219463159;
   	OWF_Key[428,9]:=1421067125;
   	OWF_Key[428,10]:=867510300;
   	OWF_Key[428,11]:=322262366;
   	OWF_Key[428,12]:=1625242888;
   	OWF_Key[428,13]:=94252119;
   	OWF_Key[428,14]:=880075177;
   	OWF_Key[428,15]:=66776100;
   	OWF_Key[428,16]:=589010987;
   	OWF_Key[429,0]:=1132727916;
   	OWF_Key[429,1]:=1932050699;
   	OWF_Key[429,2]:=2050349070;
   	OWF_Key[429,3]:=220176312;
   	OWF_Key[429,4]:=1338749261;
   	OWF_Key[429,5]:=1483219548;
   	OWF_Key[429,6]:=1142922713;
   	OWF_Key[429,7]:=652730810;
   	OWF_Key[429,8]:=1898929603;
   	OWF_Key[429,9]:=568050536;
   	OWF_Key[429,10]:=1619210705;
   	OWF_Key[429,11]:=1288733513;
   	OWF_Key[429,12]:=1326419295;
   	OWF_Key[429,13]:=980789668;
   	OWF_Key[429,14]:=2020769789;
   	OWF_Key[429,15]:=1621035431;
   	OWF_Key[429,16]:=1386884429;
   	OWF_Key[430,0]:=895139300;
   	OWF_Key[430,1]:=1724086814;
   	OWF_Key[430,2]:=930927086;
   	OWF_Key[430,3]:=1058369092;
   	OWF_Key[430,4]:=1596054800;
   	OWF_Key[430,5]:=823071432;
   	OWF_Key[430,6]:=68748739;
   	OWF_Key[430,7]:=547155910;
   	OWF_Key[430,8]:=942829868;
   	OWF_Key[430,9]:=358957743;
   	OWF_Key[430,10]:=84648904;
   	OWF_Key[430,11]:=1697774474;
   	OWF_Key[430,12]:=1084692962;
   	OWF_Key[430,13]:=2145548726;
   	OWF_Key[430,14]:=1923682716;
   	OWF_Key[430,15]:=262667437;
   	OWF_Key[430,16]:=1351416141;
   	OWF_Key[431,0]:=1114886427;
   	OWF_Key[431,1]:=438690412;
   	OWF_Key[431,2]:=202753465;
   	OWF_Key[431,3]:=1293678969;
   	OWF_Key[431,4]:=2111001365;
   	OWF_Key[431,5]:=839747077;
   	OWF_Key[431,6]:=1054397796;
   	OWF_Key[431,7]:=771999454;
   	OWF_Key[431,8]:=1111186724;
   	OWF_Key[431,9]:=1844595976;
   	OWF_Key[431,10]:=2131265084;
   	OWF_Key[431,11]:=864820484;
   	OWF_Key[431,12]:=1790775138;
   	OWF_Key[431,13]:=642693403;
   	OWF_Key[431,14]:=1450461867;
   	OWF_Key[431,15]:=2047771663;
   	OWF_Key[431,16]:=766028169;
   	OWF_Key[432,0]:=725530554;
   	OWF_Key[432,1]:=1313418696;
   	OWF_Key[432,2]:=1731227663;
   	OWF_Key[432,3]:=824223154;
   	OWF_Key[432,4]:=1232777954;
   	OWF_Key[432,5]:=1994626151;
   	OWF_Key[432,6]:=2029816048;
   	OWF_Key[432,7]:=138866526;
   	OWF_Key[432,8]:=1736142865;
   	OWF_Key[432,9]:=1872147436;
   	OWF_Key[432,10]:=689929044;
   	OWF_Key[432,11]:=2040746080;
   	OWF_Key[432,12]:=1884577054;
   	OWF_Key[432,13]:=760678168;
   	OWF_Key[432,14]:=1229480493;
   	OWF_Key[432,15]:=654878325;
   	OWF_Key[432,16]:=465908041;
   	OWF_Key[433,0]:=1802712899;
   	OWF_Key[433,1]:=469886640;
   	OWF_Key[433,2]:=1789968654;
   	OWF_Key[433,3]:=1865958582;
   	OWF_Key[433,4]:=2007611338;
   	OWF_Key[433,5]:=321976486;
   	OWF_Key[433,6]:=1263464450;
   	OWF_Key[433,7]:=829984876;
   	OWF_Key[433,8]:=1881176683;
   	OWF_Key[433,9]:=1265527937;
   	OWF_Key[433,10]:=1757714707;
   	OWF_Key[433,11]:=481681999;
   	OWF_Key[433,12]:=1169385647;
   	OWF_Key[433,13]:=1968917387;
   	OWF_Key[433,14]:=609976228;
   	OWF_Key[433,15]:=580086179;
   	OWF_Key[433,16]:=1526105979;
   	OWF_Key[434,0]:=616388254;
   	OWF_Key[434,1]:=974834252;
   	OWF_Key[434,2]:=392653343;
   	OWF_Key[434,3]:=1726973653;
   	OWF_Key[434,4]:=1824211982;
   	OWF_Key[434,5]:=1732166019;
   	OWF_Key[434,6]:=1080374198;
   	OWF_Key[434,7]:=390990230;
   	OWF_Key[434,8]:=611263632;
   	OWF_Key[434,9]:=778410222;
   	OWF_Key[434,10]:=221280023;
   	OWF_Key[434,11]:=1029717777;
   	OWF_Key[434,12]:=1445784744;
   	OWF_Key[434,13]:=1173289409;
   	OWF_Key[434,14]:=1464589909;
   	OWF_Key[434,15]:=765522900;
   	OWF_Key[434,16]:=274101697;
   	OWF_Key[435,0]:=65820213;
   	OWF_Key[435,1]:=1651646717;
   	OWF_Key[435,2]:=1786991028;
   	OWF_Key[435,3]:=1498041385;
   	OWF_Key[435,4]:=1788978986;
   	OWF_Key[435,5]:=848869242;
   	OWF_Key[435,6]:=462254383;
   	OWF_Key[435,7]:=111289191;
   	OWF_Key[435,8]:=220776889;
   	OWF_Key[435,9]:=519384734;
   	OWF_Key[435,10]:=1958864396;
   	OWF_Key[435,11]:=1812550682;
   	OWF_Key[435,12]:=1965469843;
   	OWF_Key[435,13]:=85665338;
   	OWF_Key[435,14]:=537905271;
   	OWF_Key[435,15]:=1281918993;
   	OWF_Key[435,16]:=588827800;
   	OWF_Key[436,0]:=1220204799;
   	OWF_Key[436,1]:=569892811;
   	OWF_Key[436,2]:=873297546;
   	OWF_Key[436,3]:=1409951717;
   	OWF_Key[436,4]:=373999743;
   	OWF_Key[436,5]:=955795349;
   	OWF_Key[436,6]:=1056576480;
   	OWF_Key[436,7]:=2093776834;
   	OWF_Key[436,8]:=504508589;